VERSION : 0.1
// Master sequencing for automatic operation
   VAR_INPUT
      RST : Bool;   // Sequence reset
   END_VAR
   VAR_OUTPUT
      RNG : Bool;   // Sequence running
   END_VAR
   VAR
      CRNT_STEP : Int;
      STEP_001 : "500_SEQ_STEP";
      STEP_005 : "500_SEQ_STEP";
      STEP_010 : "500_SEQ_STEP";
      STEP_020 : "500_SEQ_STEP";
      STEP_030 : "500_SEQ_STEP";
      STEP_040 : "500_SEQ_STEP";
      STEP_050 : "500_SEQ_STEP";
      STEP_060 : "500_SEQ_STEP";
      STEP_070 : "500_SEQ_STEP";
      STEP_080 : "500_SEQ_STEP";
      STEP_090 : "500_SEQ_STEP";
      STEP_095 : "500_SEQ_STEP";
      STEP_100 : "500_SEQ_STEP";
      STEP_110 : "500_SEQ_STEP";
      STEP_120 : "500_SEQ_STEP";
      STEP_130 : "500_SEQ_STEP";
      STEP_140 : "500_SEQ_STEP";
      STEP_150 : "500_SEQ_STEP";
      STEP_160 : "500_SEQ_STEP";
      STEP_170 : "500_SEQ_STEP";
      STEP_180 : "500_SEQ_STEP";
      STEP_190 : "500_SEQ_STEP";
      STEP_200 : "500_SEQ_STEP";
      STEP_210 : "500_SEQ_STEP";
      STEP_220 : "500_SEQ_STEP";
      STEP_230 : "500_SEQ_STEP";
      STEP_240 : "500_SEQ_STEP";
      STEP_250 : "500_SEQ_STEP";
      STEP_260 : "500_SEQ_STEP";
      STEP_270 : "500_SEQ_STEP";
      STEP_300 : "500_SEQ_STEP";
      STEP_310 : "500_SEQ_STEP";
      STEP_320 : "500_SEQ_STEP";
      STEP_330 : "500_SEQ_STEP";
      STEP_340 : "500_SEQ_STEP";
      STEP_350 : "500_SEQ_STEP";
      STEP_360 : "500_SEQ_STEP";
      STEP_370 : "500_SEQ_STEP";
      STEP_380 : "500_SEQ_STEP";
      STEP_390 : "500_SEQ_STEP";
      STEP_400 : "500_SEQ_STEP";
      STEP_410 : "500_SEQ_STEP";
      STEP_420 : "500_SEQ_STEP";
      STEP_430 : "500_SEQ_STEP";
      STEP_440 : "500_SEQ_STEP";
      STEP_450 : "500_SEQ_STEP";
      STEP_460 : "500_SEQ_STEP";
      STEP_470 : "500_SEQ_STEP";
      STEP_480 : "500_SEQ_STEP";
      STEP_490 : "500_SEQ_STEP";
      STEP_500 : "500_SEQ_STEP";
      STEP_510 : "500_SEQ_STEP";
      STEP_520 : "500_SEQ_STEP";
      STEP_525 : "500_SEQ_STEP";
      STEP_530 : "500_SEQ_STEP";
      STEP_540 : "500_SEQ_STEP";
      STEP_550 : "500_SEQ_STEP";
      STEP_560 : "500_SEQ_STEP";
      STEP_570 : "500_SEQ_STEP";
   END_VAR
   VAR_TEMP   // added for the SCL form of the ladder/FBD networks
      _w1 : Bool;
   END_VAR
BEGIN

REGION Network 1: Auto Initiated or Reset = Set Step to 0
   // Going into automatic or sequence reset resets the sequence
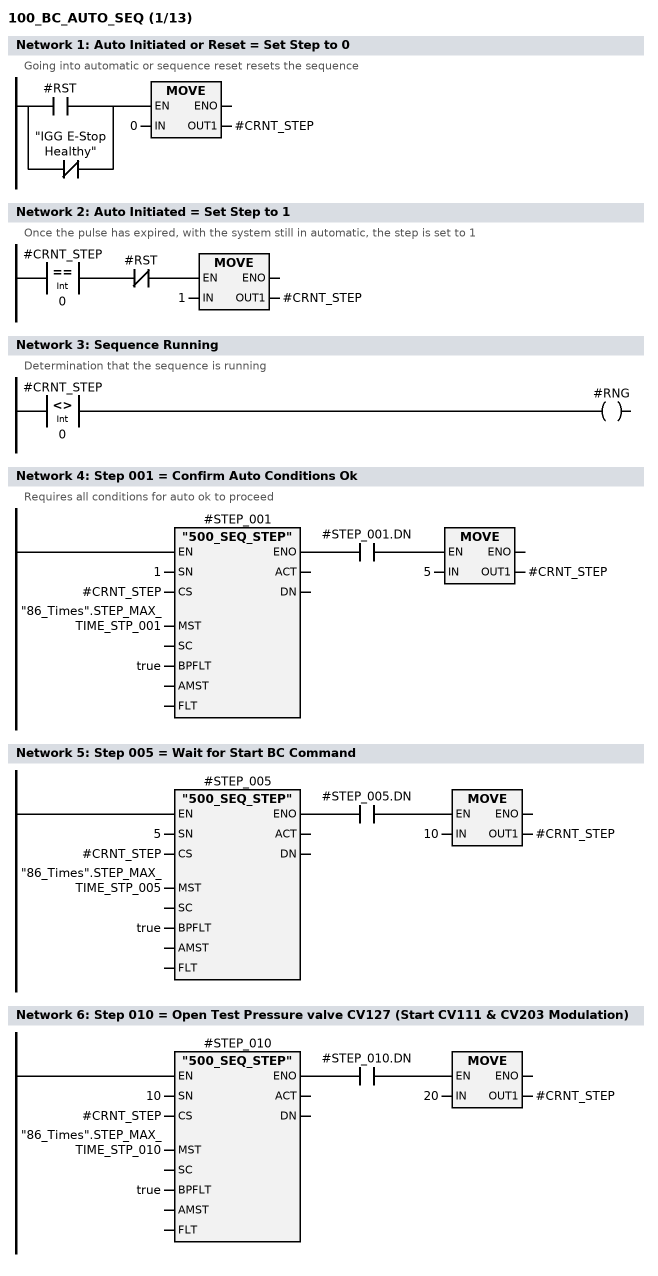
   RUNG wire#powerrail
      Contact( #RST )
      wire#w1
      Move(in := 0, out1 => #CRNT_STEP)
   END_RUNG
   RUNG wire#powerrail
      I_Contact( "IGG E-Stop Healthy" )
   END_RUNG wire#w1
   // the same network as SCL:
   IF #RST OR NOT "IGG E-Stop Healthy" THEN #CRNT_STEP := 0; END_IF;
END_REGION

REGION Network 2: Auto Initiated = Set Step to 1
   // Once the pulse has expired, with the system still in automatic, the step is set to 1
   RUNG wire#powerrail
      { S7_Templates := "SrcType := Int" } EQ_Contact(in1 := #CRNT_STEP, in2 := 0)
      I_Contact( #RST )
      Move(in := 1, out1 => #CRNT_STEP)
   END_RUNG
   // the same network as SCL:
   IF (#CRNT_STEP = 0) AND NOT #RST THEN #CRNT_STEP := 1; END_IF;
END_REGION

REGION Network 3: Sequence Running
   // Determination that the sequence is running
   RUNG wire#powerrail
      { S7_Templates := "SrcType := Int" } NE_Contact(in1 := #CRNT_STEP, in2 := 0)
      Coil( #RNG )
   END_RUNG
   // the same network as SCL:
   #RNG := #CRNT_STEP <> 0;
END_REGION

REGION Network 4: Step 001 = Confirm Auto Conditions Ok
   // Requires all conditions for auto ok to proceed
   RUNG wire#powerrail
      #STEP_001(SN := 1, CS := #CRNT_STEP, MST := "86_Times".STEP_MAX_TIME_STP_001, SC :=, BPFLT := true, AMST :=, FLT :=, ACT =>, DN =>)
      Contact( #STEP_001.DN )
      Move(in := 5, out1 => #CRNT_STEP)
   END_RUNG
   // the same network as SCL:
   #STEP_001(SN := 1, CS := #CRNT_STEP, MST := "86_Times".STEP_MAX_TIME_STP_001, BPFLT := true, ENO => #_w1);   // "500_SEQ_STEP"
   IF #_w1 AND #STEP_001.DN THEN #CRNT_STEP := 5; END_IF;
END_REGION

REGION Network 5: Step 005 = Wait for Start BC Command
   RUNG wire#powerrail
      #STEP_005(SN := 5, CS := #CRNT_STEP, MST := "86_Times".STEP_MAX_TIME_STP_005, SC :=, BPFLT := true, AMST :=, FLT :=, ACT =>, DN =>)
      Contact( #STEP_005.DN )
      Move(in := 10, out1 => #CRNT_STEP)
   END_RUNG
   // the same network as SCL:
   #STEP_005(SN := 5, CS := #CRNT_STEP, MST := "86_Times".STEP_MAX_TIME_STP_005, BPFLT := true, ENO => #_w1);   // "500_SEQ_STEP"
   IF #_w1 AND #STEP_005.DN THEN #CRNT_STEP := 10; END_IF;
END_REGION

REGION Network 6: Step 010 = Open Test Pressure valve CV127 (Start CV111 & CV203 Modulation)
   RUNG wire#powerrail
      #STEP_010(SN := 10, CS := #CRNT_STEP, MST := "86_Times".STEP_MAX_TIME_STP_010, SC :=, BPFLT := true, AMST :=, FLT :=, ACT =>, DN =>)
      Contact( #STEP_010.DN )
      Move(in := 20, out1 => #CRNT_STEP)
   END_RUNG
   // the same network as SCL:
   #STEP_010(SN := 10, CS := #CRNT_STEP, MST := "86_Times".STEP_MAX_TIME_STP_010, BPFLT := true, ENO => #_w1);   // "500_SEQ_STEP"
   IF #_w1 AND #STEP_010.DN THEN #CRNT_STEP := 20; END_IF;
END_REGION

REGION Network 7: Step 020 = Check Pressure PS101
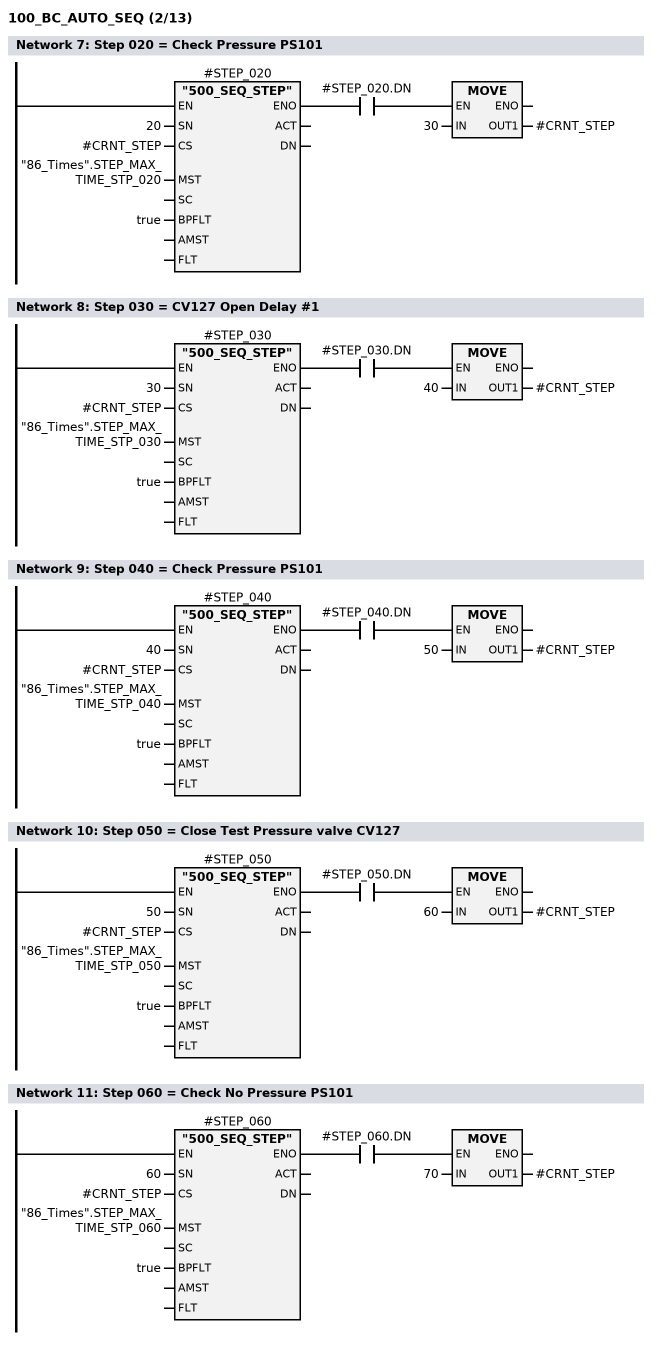
   RUNG wire#powerrail
      #STEP_020(SN := 20, CS := #CRNT_STEP, MST := "86_Times".STEP_MAX_TIME_STP_020, SC :=, BPFLT := true, AMST :=, FLT :=, ACT =>, DN =>)
      Contact( #STEP_020.DN )
      Move(in := 30, out1 => #CRNT_STEP)
   END_RUNG
   // the same network as SCL:
   #STEP_020(SN := 20, CS := #CRNT_STEP, MST := "86_Times".STEP_MAX_TIME_STP_020, BPFLT := true, ENO => #_w1);   // "500_SEQ_STEP"
   IF #_w1 AND #STEP_020.DN THEN #CRNT_STEP := 30; END_IF;
END_REGION

REGION Network 8: Step 030 = CV127 Open Delay #1
   RUNG wire#powerrail
      #STEP_030(SN := 30, CS := #CRNT_STEP, MST := "86_Times".STEP_MAX_TIME_STP_030, SC :=, BPFLT := true, AMST :=, FLT :=, ACT =>, DN =>)
      Contact( #STEP_030.DN )
      Move(in := 40, out1 => #CRNT_STEP)
   END_RUNG
   // the same network as SCL:
   #STEP_030(SN := 30, CS := #CRNT_STEP, MST := "86_Times".STEP_MAX_TIME_STP_030, BPFLT := true, ENO => #_w1);   // "500_SEQ_STEP"
   IF #_w1 AND #STEP_030.DN THEN #CRNT_STEP := 40; END_IF;
END_REGION

REGION Network 9: Step 040 = Check Pressure PS101
   RUNG wire#powerrail
      #STEP_040(SN := 40, CS := #CRNT_STEP, MST := "86_Times".STEP_MAX_TIME_STP_040, SC :=, BPFLT := true, AMST :=, FLT :=, ACT =>, DN =>)
      Contact( #STEP_040.DN )
      Move(in := 50, out1 => #CRNT_STEP)
   END_RUNG
   // the same network as SCL:
   #STEP_040(SN := 40, CS := #CRNT_STEP, MST := "86_Times".STEP_MAX_TIME_STP_040, BPFLT := true, ENO => #_w1);   // "500_SEQ_STEP"
   IF #_w1 AND #STEP_040.DN THEN #CRNT_STEP := 50; END_IF;
END_REGION

REGION Network 10: Step 050 = Close Test Pressure valve CV127
   RUNG wire#powerrail
      #STEP_050(SN := 50, CS := #CRNT_STEP, MST := "86_Times".STEP_MAX_TIME_STP_050, SC :=, BPFLT := true, AMST :=, FLT :=, ACT =>, DN =>)
      Contact( #STEP_050.DN )
      Move(in := 60, out1 => #CRNT_STEP)
   END_RUNG
   // the same network as SCL:
   #STEP_050(SN := 50, CS := #CRNT_STEP, MST := "86_Times".STEP_MAX_TIME_STP_050, BPFLT := true, ENO => #_w1);   // "500_SEQ_STEP"
   IF #_w1 AND #STEP_050.DN THEN #CRNT_STEP := 60; END_IF;
END_REGION

REGION Network 11: Step 060 = Check No Pressure PS101
   RUNG wire#powerrail
      #STEP_060(SN := 60, CS := #CRNT_STEP, MST := "86_Times".STEP_MAX_TIME_STP_060, SC :=, BPFLT := true, AMST :=, FLT :=, ACT =>, DN =>)
      Contact( #STEP_060.DN )
      Move(in := 70, out1 => #CRNT_STEP)
   END_RUNG
   // the same network as SCL:
   #STEP_060(SN := 60, CS := #CRNT_STEP, MST := "86_Times".STEP_MAX_TIME_STP_060, BPFLT := true, ENO => #_w1);   // "500_SEQ_STEP"
   IF #_w1 AND #STEP_060.DN THEN #CRNT_STEP := 70; END_IF;
END_REGION

REGION Network 12: Step 070 = CV127 Closed Delay
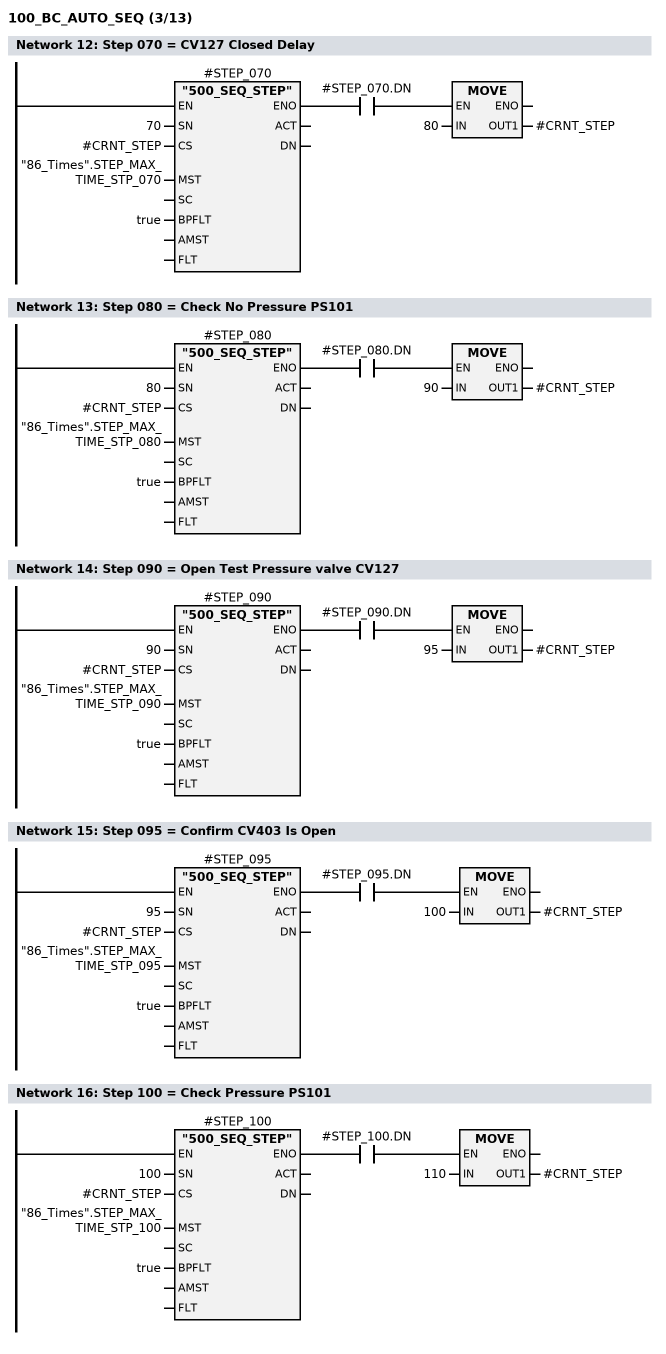
   RUNG wire#powerrail
      #STEP_070(SN := 70, CS := #CRNT_STEP, MST := "86_Times".STEP_MAX_TIME_STP_070, SC :=, BPFLT := true, AMST :=, FLT :=, ACT =>, DN =>)
      Contact( #STEP_070.DN )
      Move(in := 80, out1 => #CRNT_STEP)
   END_RUNG
   // the same network as SCL:
   #STEP_070(SN := 70, CS := #CRNT_STEP, MST := "86_Times".STEP_MAX_TIME_STP_070, BPFLT := true, ENO => #_w1);   // "500_SEQ_STEP"
   IF #_w1 AND #STEP_070.DN THEN #CRNT_STEP := 80; END_IF;
END_REGION

REGION Network 13: Step 080 = Check No Pressure PS101
   RUNG wire#powerrail
      #STEP_080(SN := 80, CS := #CRNT_STEP, MST := "86_Times".STEP_MAX_TIME_STP_080, SC :=, BPFLT := true, AMST :=, FLT :=, ACT =>, DN =>)
      Contact( #STEP_080.DN )
      Move(in := 90, out1 => #CRNT_STEP)
   END_RUNG
   // the same network as SCL:
   #STEP_080(SN := 80, CS := #CRNT_STEP, MST := "86_Times".STEP_MAX_TIME_STP_080, BPFLT := true, ENO => #_w1);   // "500_SEQ_STEP"
   IF #_w1 AND #STEP_080.DN THEN #CRNT_STEP := 90; END_IF;
END_REGION

REGION Network 14: Step 090 = Open Test Pressure valve CV127
   RUNG wire#powerrail
      #STEP_090(SN := 90, CS := #CRNT_STEP, MST := "86_Times".STEP_MAX_TIME_STP_090, SC :=, BPFLT := true, AMST :=, FLT :=, ACT =>, DN =>)
      Contact( #STEP_090.DN )
      Move(in := 95, out1 => #CRNT_STEP)
   END_RUNG
   // the same network as SCL:
   #STEP_090(SN := 90, CS := #CRNT_STEP, MST := "86_Times".STEP_MAX_TIME_STP_090, BPFLT := true, ENO => #_w1);   // "500_SEQ_STEP"
   IF #_w1 AND #STEP_090.DN THEN #CRNT_STEP := 95; END_IF;
END_REGION

REGION Network 15: Step 095 = Confirm CV403 Is Open
   RUNG wire#powerrail
      #STEP_095(SN := 95, CS := #CRNT_STEP, MST := "86_Times".STEP_MAX_TIME_STP_095, SC :=, BPFLT := true, AMST :=, FLT :=, ACT =>, DN =>)
      Contact( #STEP_095.DN )
      Move(in := 100, out1 => #CRNT_STEP)
   END_RUNG
   // the same network as SCL:
   #STEP_095(SN := 95, CS := #CRNT_STEP, MST := "86_Times".STEP_MAX_TIME_STP_095, BPFLT := true, ENO => #_w1);   // "500_SEQ_STEP"
   IF #_w1 AND #STEP_095.DN THEN #CRNT_STEP := 100; END_IF;
END_REGION

REGION Network 16: Step 100 = Check Pressure PS101
   RUNG wire#powerrail
      #STEP_100(SN := 100, CS := #CRNT_STEP, MST := "86_Times".STEP_MAX_TIME_STP_100, SC :=, BPFLT := true, AMST :=, FLT :=, ACT =>, DN =>)
      Contact( #STEP_100.DN )
      Move(in := 110, out1 => #CRNT_STEP)
   END_RUNG
   // the same network as SCL:
   #STEP_100(SN := 100, CS := #CRNT_STEP, MST := "86_Times".STEP_MAX_TIME_STP_100, BPFLT := true, ENO => #_w1);   // "500_SEQ_STEP"
   IF #_w1 AND #STEP_100.DN THEN #CRNT_STEP := 110; END_IF;
END_REGION

REGION Network 17: Step110 = CV127 Open Delay #2
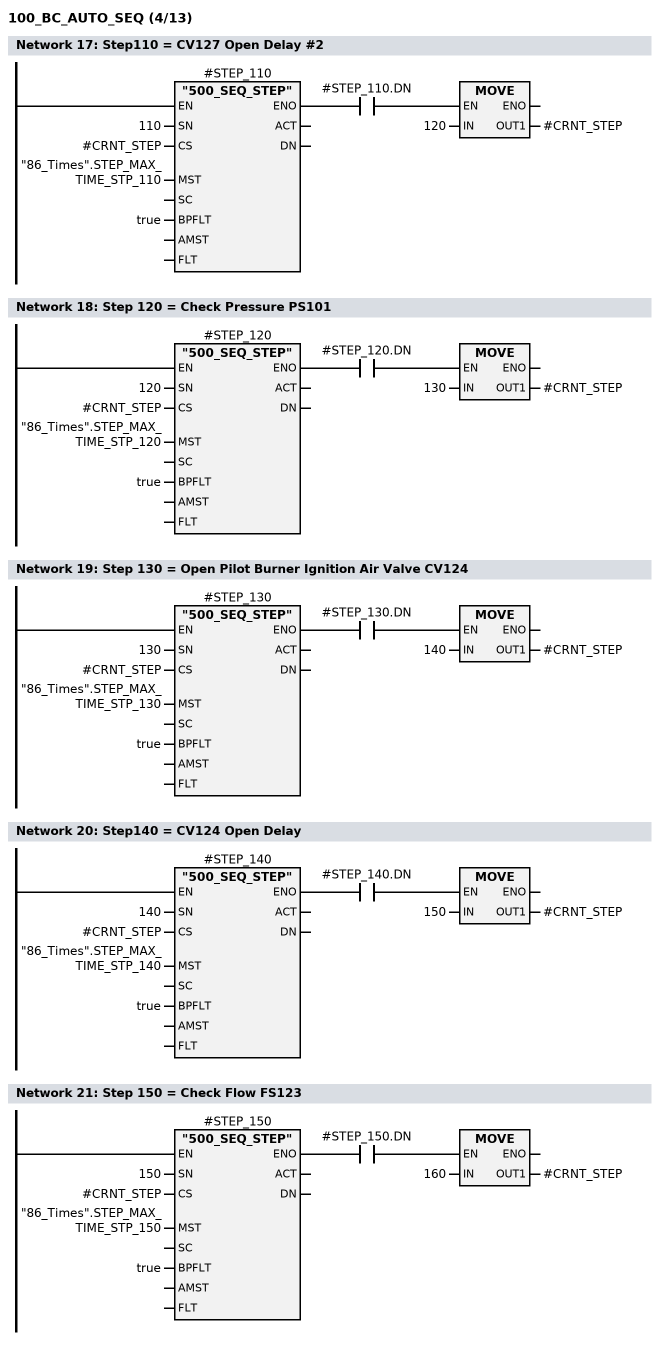
   RUNG wire#powerrail
      #STEP_110(SN := 110, CS := #CRNT_STEP, MST := "86_Times".STEP_MAX_TIME_STP_110, SC :=, BPFLT := true, AMST :=, FLT :=, ACT =>, DN =>)
      Contact( #STEP_110.DN )
      Move(in := 120, out1 => #CRNT_STEP)
   END_RUNG
   // the same network as SCL:
   #STEP_110(SN := 110, CS := #CRNT_STEP, MST := "86_Times".STEP_MAX_TIME_STP_110, BPFLT := true, ENO => #_w1);   // "500_SEQ_STEP"
   IF #_w1 AND #STEP_110.DN THEN #CRNT_STEP := 120; END_IF;
END_REGION

REGION Network 18: Step 120 = Check Pressure PS101
   RUNG wire#powerrail
      #STEP_120(SN := 120, CS := #CRNT_STEP, MST := "86_Times".STEP_MAX_TIME_STP_120, SC :=, BPFLT := true, AMST :=, FLT :=, ACT =>, DN =>)
      Contact( #STEP_120.DN )
      Move(in := 130, out1 => #CRNT_STEP)
   END_RUNG
   // the same network as SCL:
   #STEP_120(SN := 120, CS := #CRNT_STEP, MST := "86_Times".STEP_MAX_TIME_STP_120, BPFLT := true, ENO => #_w1);   // "500_SEQ_STEP"
   IF #_w1 AND #STEP_120.DN THEN #CRNT_STEP := 130; END_IF;
END_REGION

REGION Network 19: Step 130 = Open Pilot Burner Ignition Air Valve CV124
   RUNG wire#powerrail
      #STEP_130(SN := 130, CS := #CRNT_STEP, MST := "86_Times".STEP_MAX_TIME_STP_130, SC :=, BPFLT := true, AMST :=, FLT :=, ACT =>, DN =>)
      Contact( #STEP_130.DN )
      Move(in := 140, out1 => #CRNT_STEP)
   END_RUNG
   // the same network as SCL:
   #STEP_130(SN := 130, CS := #CRNT_STEP, MST := "86_Times".STEP_MAX_TIME_STP_130, BPFLT := true, ENO => #_w1);   // "500_SEQ_STEP"
   IF #_w1 AND #STEP_130.DN THEN #CRNT_STEP := 140; END_IF;
END_REGION

REGION Network 20: Step140 = CV124 Open Delay
   RUNG wire#powerrail
      #STEP_140(SN := 140, CS := #CRNT_STEP, MST := "86_Times".STEP_MAX_TIME_STP_140, SC :=, BPFLT := true, AMST :=, FLT :=, ACT =>, DN =>)
      Contact( #STEP_140.DN )
      Move(in := 150, out1 => #CRNT_STEP)
   END_RUNG
   // the same network as SCL:
   #STEP_140(SN := 140, CS := #CRNT_STEP, MST := "86_Times".STEP_MAX_TIME_STP_140, BPFLT := true, ENO => #_w1);   // "500_SEQ_STEP"
   IF #_w1 AND #STEP_140.DN THEN #CRNT_STEP := 150; END_IF;
END_REGION

REGION Network 21: Step 150 = Check Flow FS123
   RUNG wire#powerrail
      #STEP_150(SN := 150, CS := #CRNT_STEP, MST := "86_Times".STEP_MAX_TIME_STP_150, SC :=, BPFLT := true, AMST :=, FLT :=, ACT =>, DN =>)
      Contact( #STEP_150.DN )
      Move(in := 160, out1 => #CRNT_STEP)
   END_RUNG
   // the same network as SCL:
   #STEP_150(SN := 150, CS := #CRNT_STEP, MST := "86_Times".STEP_MAX_TIME_STP_150, BPFLT := true, ENO => #_w1);   // "500_SEQ_STEP"
   IF #_w1 AND #STEP_150.DN THEN #CRNT_STEP := 160; END_IF;
END_REGION

REGION Network 22: Step 160 = Pilot Flame Ignition Sequence
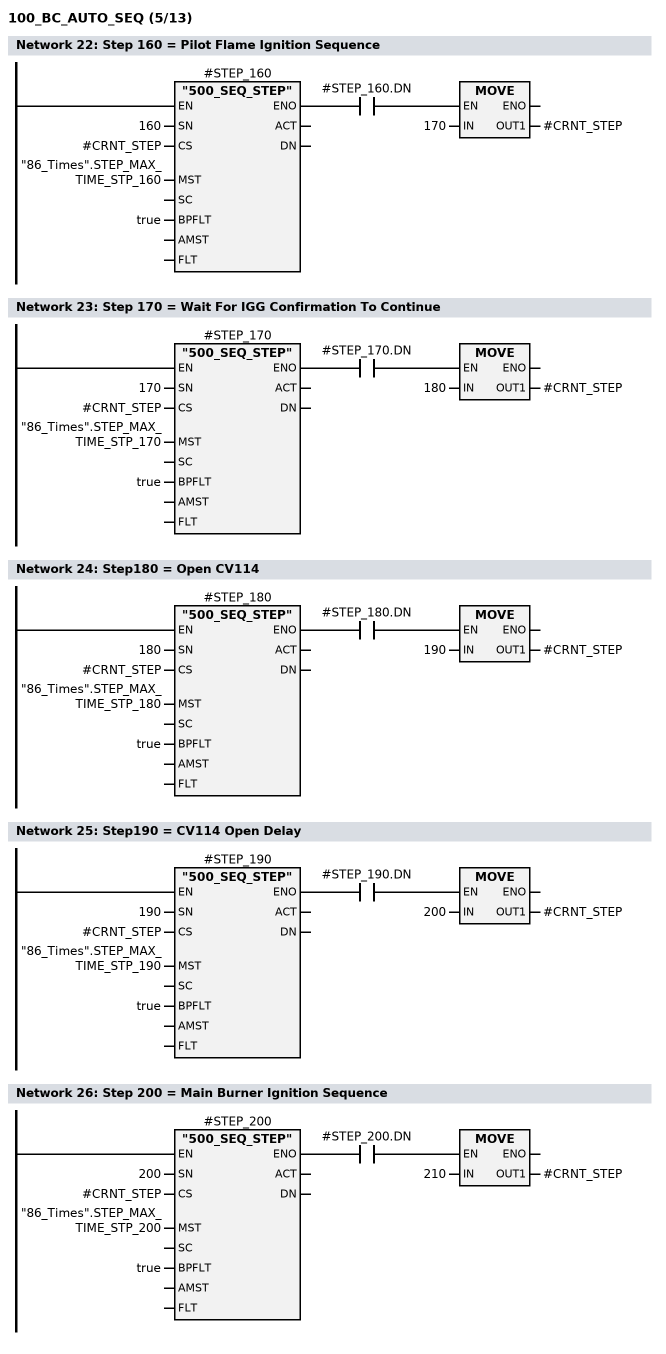
   RUNG wire#powerrail
      #STEP_160(SN := 160, CS := #CRNT_STEP, MST := "86_Times".STEP_MAX_TIME_STP_160, SC :=, BPFLT := true, AMST :=, FLT :=, ACT =>, DN =>)
      Contact( #STEP_160.DN )
      Move(in := 170, out1 => #CRNT_STEP)
   END_RUNG
   // the same network as SCL:
   #STEP_160(SN := 160, CS := #CRNT_STEP, MST := "86_Times".STEP_MAX_TIME_STP_160, BPFLT := true, ENO => #_w1);   // "500_SEQ_STEP"
   IF #_w1 AND #STEP_160.DN THEN #CRNT_STEP := 170; END_IF;
END_REGION

REGION Network 23: Step 170 = Wait For IGG Confirmation To Continue
   RUNG wire#powerrail
      #STEP_170(SN := 170, CS := #CRNT_STEP, MST := "86_Times".STEP_MAX_TIME_STP_170, SC :=, BPFLT := true, AMST :=, FLT :=, ACT =>, DN =>)
      Contact( #STEP_170.DN )
      Move(in := 180, out1 => #CRNT_STEP)
   END_RUNG
   // the same network as SCL:
   #STEP_170(SN := 170, CS := #CRNT_STEP, MST := "86_Times".STEP_MAX_TIME_STP_170, BPFLT := true, ENO => #_w1);   // "500_SEQ_STEP"
   IF #_w1 AND #STEP_170.DN THEN #CRNT_STEP := 180; END_IF;
END_REGION

REGION Network 24: Step180 = Open CV114
   RUNG wire#powerrail
      #STEP_180(SN := 180, CS := #CRNT_STEP, MST := "86_Times".STEP_MAX_TIME_STP_180, SC :=, BPFLT := true, AMST :=, FLT :=, ACT =>, DN =>)
      Contact( #STEP_180.DN )
      Move(in := 190, out1 => #CRNT_STEP)
   END_RUNG
   // the same network as SCL:
   #STEP_180(SN := 180, CS := #CRNT_STEP, MST := "86_Times".STEP_MAX_TIME_STP_180, BPFLT := true, ENO => #_w1);   // "500_SEQ_STEP"
   IF #_w1 AND #STEP_180.DN THEN #CRNT_STEP := 190; END_IF;
END_REGION

REGION Network 25: Step190 = CV114 Open Delay
   RUNG wire#powerrail
      #STEP_190(SN := 190, CS := #CRNT_STEP, MST := "86_Times".STEP_MAX_TIME_STP_190, SC :=, BPFLT := true, AMST :=, FLT :=, ACT =>, DN =>)
      Contact( #STEP_190.DN )
      Move(in := 200, out1 => #CRNT_STEP)
   END_RUNG
   // the same network as SCL:
   #STEP_190(SN := 190, CS := #CRNT_STEP, MST := "86_Times".STEP_MAX_TIME_STP_190, BPFLT := true, ENO => #_w1);   // "500_SEQ_STEP"
   IF #_w1 AND #STEP_190.DN THEN #CRNT_STEP := 200; END_IF;
END_REGION

REGION Network 26: Step 200 = Main Burner Ignition Sequence
   RUNG wire#powerrail
      #STEP_200(SN := 200, CS := #CRNT_STEP, MST := "86_Times".STEP_MAX_TIME_STP_200, SC :=, BPFLT := true, AMST :=, FLT :=, ACT =>, DN =>)
      Contact( #STEP_200.DN )
      Move(in := 210, out1 => #CRNT_STEP)
   END_RUNG
   // the same network as SCL:
   #STEP_200(SN := 200, CS := #CRNT_STEP, MST := "86_Times".STEP_MAX_TIME_STP_200, BPFLT := true, ENO => #_w1);   // "500_SEQ_STEP"
   IF #_w1 AND #STEP_200.DN THEN #CRNT_STEP := 210; END_IF;
END_REGION

REGION Network 27: Step 210 = Check Pressure PIT113
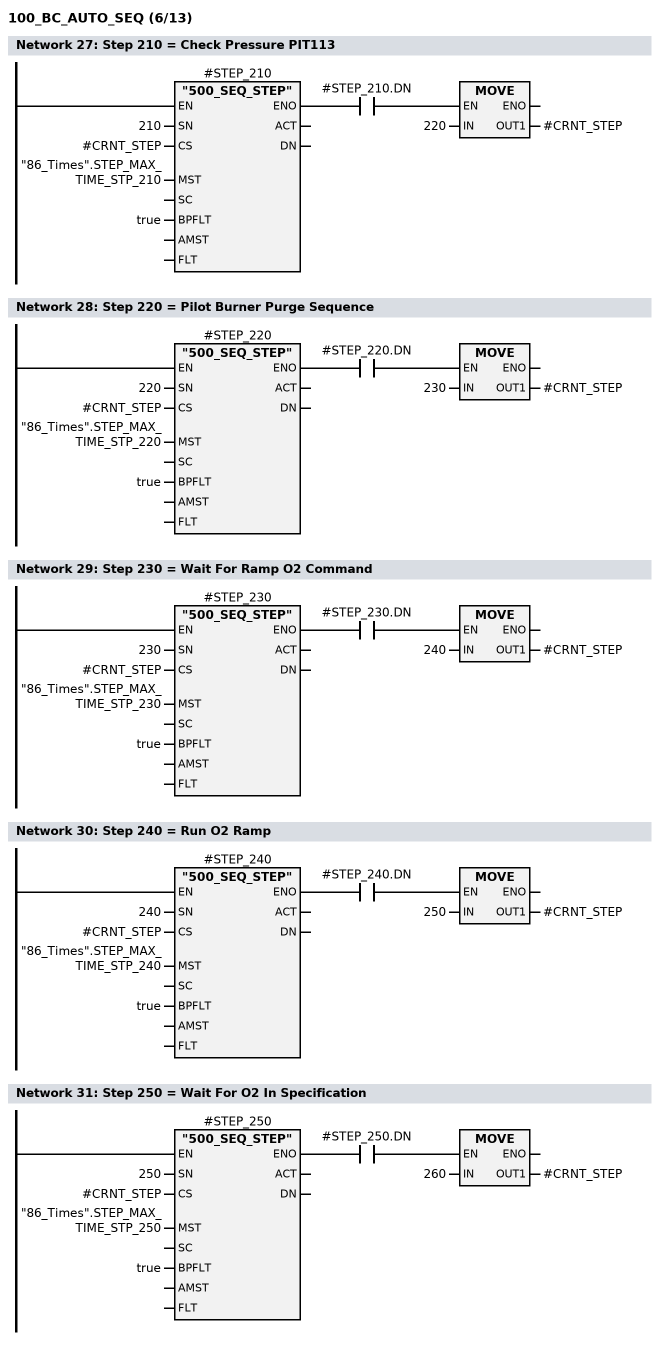
   RUNG wire#powerrail
      #STEP_210(SN := 210, CS := #CRNT_STEP, MST := "86_Times".STEP_MAX_TIME_STP_210, SC :=, BPFLT := true, AMST :=, FLT :=, ACT =>, DN =>)
      Contact( #STEP_210.DN )
      Move(in := 220, out1 => #CRNT_STEP)
   END_RUNG
   // the same network as SCL:
   #STEP_210(SN := 210, CS := #CRNT_STEP, MST := "86_Times".STEP_MAX_TIME_STP_210, BPFLT := true, ENO => #_w1);   // "500_SEQ_STEP"
   IF #_w1 AND #STEP_210.DN THEN #CRNT_STEP := 220; END_IF;
END_REGION

REGION Network 28: Step 220 = Pilot Burner Purge Sequence
   RUNG wire#powerrail
      #STEP_220(SN := 220, CS := #CRNT_STEP, MST := "86_Times".STEP_MAX_TIME_STP_220, SC :=, BPFLT := true, AMST :=, FLT :=, ACT =>, DN =>)
      Contact( #STEP_220.DN )
      Move(in := 230, out1 => #CRNT_STEP)
   END_RUNG
   // the same network as SCL:
   #STEP_220(SN := 220, CS := #CRNT_STEP, MST := "86_Times".STEP_MAX_TIME_STP_220, BPFLT := true, ENO => #_w1);   // "500_SEQ_STEP"
   IF #_w1 AND #STEP_220.DN THEN #CRNT_STEP := 230; END_IF;
END_REGION

REGION Network 29: Step 230 = Wait For Ramp O2 Command
   RUNG wire#powerrail
      #STEP_230(SN := 230, CS := #CRNT_STEP, MST := "86_Times".STEP_MAX_TIME_STP_230, SC :=, BPFLT := true, AMST :=, FLT :=, ACT =>, DN =>)
      Contact( #STEP_230.DN )
      Move(in := 240, out1 => #CRNT_STEP)
   END_RUNG
   // the same network as SCL:
   #STEP_230(SN := 230, CS := #CRNT_STEP, MST := "86_Times".STEP_MAX_TIME_STP_230, BPFLT := true, ENO => #_w1);   // "500_SEQ_STEP"
   IF #_w1 AND #STEP_230.DN THEN #CRNT_STEP := 240; END_IF;
END_REGION

REGION Network 30: Step 240 = Run O2 Ramp
   RUNG wire#powerrail
      #STEP_240(SN := 240, CS := #CRNT_STEP, MST := "86_Times".STEP_MAX_TIME_STP_240, SC :=, BPFLT := true, AMST :=, FLT :=, ACT =>, DN =>)
      Contact( #STEP_240.DN )
      Move(in := 250, out1 => #CRNT_STEP)
   END_RUNG
   // the same network as SCL:
   #STEP_240(SN := 240, CS := #CRNT_STEP, MST := "86_Times".STEP_MAX_TIME_STP_240, BPFLT := true, ENO => #_w1);   // "500_SEQ_STEP"
   IF #_w1 AND #STEP_240.DN THEN #CRNT_STEP := 250; END_IF;
END_REGION

REGION Network 31: Step 250 = Wait For O2 In Specification
   RUNG wire#powerrail
      #STEP_250(SN := 250, CS := #CRNT_STEP, MST := "86_Times".STEP_MAX_TIME_STP_250, SC :=, BPFLT := true, AMST :=, FLT :=, ACT =>, DN =>)
      Contact( #STEP_250.DN )
      Move(in := 260, out1 => #CRNT_STEP)
   END_RUNG
   // the same network as SCL:
   #STEP_250(SN := 250, CS := #CRNT_STEP, MST := "86_Times".STEP_MAX_TIME_STP_250, BPFLT := true, ENO => #_w1);   // "500_SEQ_STEP"
   IF #_w1 AND #STEP_250.DN THEN #CRNT_STEP := 260; END_IF;
END_REGION

REGION Network 32: Step 260 = Write O2 Within Specification Status To IGG
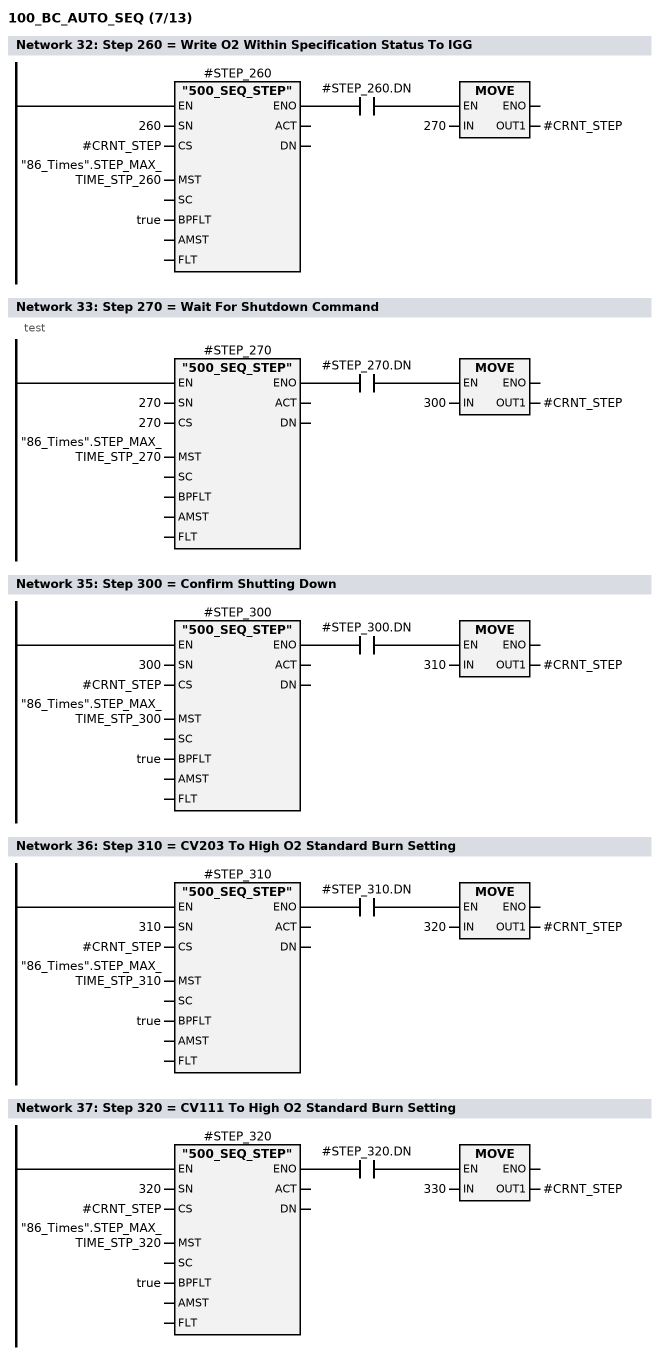
   RUNG wire#powerrail
      #STEP_260(SN := 260, CS := #CRNT_STEP, MST := "86_Times".STEP_MAX_TIME_STP_260, SC :=, BPFLT := true, AMST :=, FLT :=, ACT =>, DN =>)
      Contact( #STEP_260.DN )
      Move(in := 270, out1 => #CRNT_STEP)
   END_RUNG
   // the same network as SCL:
   #STEP_260(SN := 260, CS := #CRNT_STEP, MST := "86_Times".STEP_MAX_TIME_STP_260, BPFLT := true, ENO => #_w1);   // "500_SEQ_STEP"
   IF #_w1 AND #STEP_260.DN THEN #CRNT_STEP := 270; END_IF;
END_REGION

REGION Network 33: Step 270 = Wait For Shutdown Command
   // test
   RUNG wire#powerrail
      #STEP_270(SN := 270, CS := 270, MST := "86_Times".STEP_MAX_TIME_STP_270, SC :=, BPFLT :=, AMST :=, FLT :=, ACT =>, DN =>)
      Contact( #STEP_270.DN )
      Move(in := 300, out1 => #CRNT_STEP)
   END_RUNG
   // the same network as SCL:
   #STEP_270(SN := 270, CS := 270, MST := "86_Times".STEP_MAX_TIME_STP_270, ENO => #_w1);   // "500_SEQ_STEP"
   IF #_w1 AND #STEP_270.DN THEN #CRNT_STEP := 300; END_IF;
END_REGION

REGION Network 35: Step 300 = Confirm Shutting Down
   RUNG wire#powerrail
      #STEP_300(SN := 300, CS := #CRNT_STEP, MST := "86_Times".STEP_MAX_TIME_STP_300, SC :=, BPFLT := true, AMST :=, FLT :=, ACT =>, DN =>)
      Contact( #STEP_300.DN )
      Move(in := 310, out1 => #CRNT_STEP)
   END_RUNG
   // the same network as SCL:
   #STEP_300(SN := 300, CS := #CRNT_STEP, MST := "86_Times".STEP_MAX_TIME_STP_300, BPFLT := true, ENO => #_w1);   // "500_SEQ_STEP"
   IF #_w1 AND #STEP_300.DN THEN #CRNT_STEP := 310; END_IF;
END_REGION

REGION Network 36: Step 310 = CV203 To High O2 Standard Burn Setting
   RUNG wire#powerrail
      #STEP_310(SN := 310, CS := #CRNT_STEP, MST := "86_Times".STEP_MAX_TIME_STP_310, SC :=, BPFLT := true, AMST :=, FLT :=, ACT =>, DN =>)
      Contact( #STEP_310.DN )
      Move(in := 320, out1 => #CRNT_STEP)
   END_RUNG
   // the same network as SCL:
   #STEP_310(SN := 310, CS := #CRNT_STEP, MST := "86_Times".STEP_MAX_TIME_STP_310, BPFLT := true, ENO => #_w1);   // "500_SEQ_STEP"
   IF #_w1 AND #STEP_310.DN THEN #CRNT_STEP := 320; END_IF;
END_REGION

REGION Network 37: Step 320 = CV111 To High O2 Standard Burn Setting
   RUNG wire#powerrail
      #STEP_320(SN := 320, CS := #CRNT_STEP, MST := "86_Times".STEP_MAX_TIME_STP_320, SC :=, BPFLT := true, AMST :=, FLT :=, ACT =>, DN =>)
      Contact( #STEP_320.DN )
      Move(in := 330, out1 => #CRNT_STEP)
   END_RUNG
   // the same network as SCL:
   #STEP_320(SN := 320, CS := #CRNT_STEP, MST := "86_Times".STEP_MAX_TIME_STP_320, BPFLT := true, ENO => #_w1);   // "500_SEQ_STEP"
   IF #_w1 AND #STEP_320.DN THEN #CRNT_STEP := 330; END_IF;
END_REGION

REGION Network 38: Step 330 = Modulation Stopped Confirmation To IGG
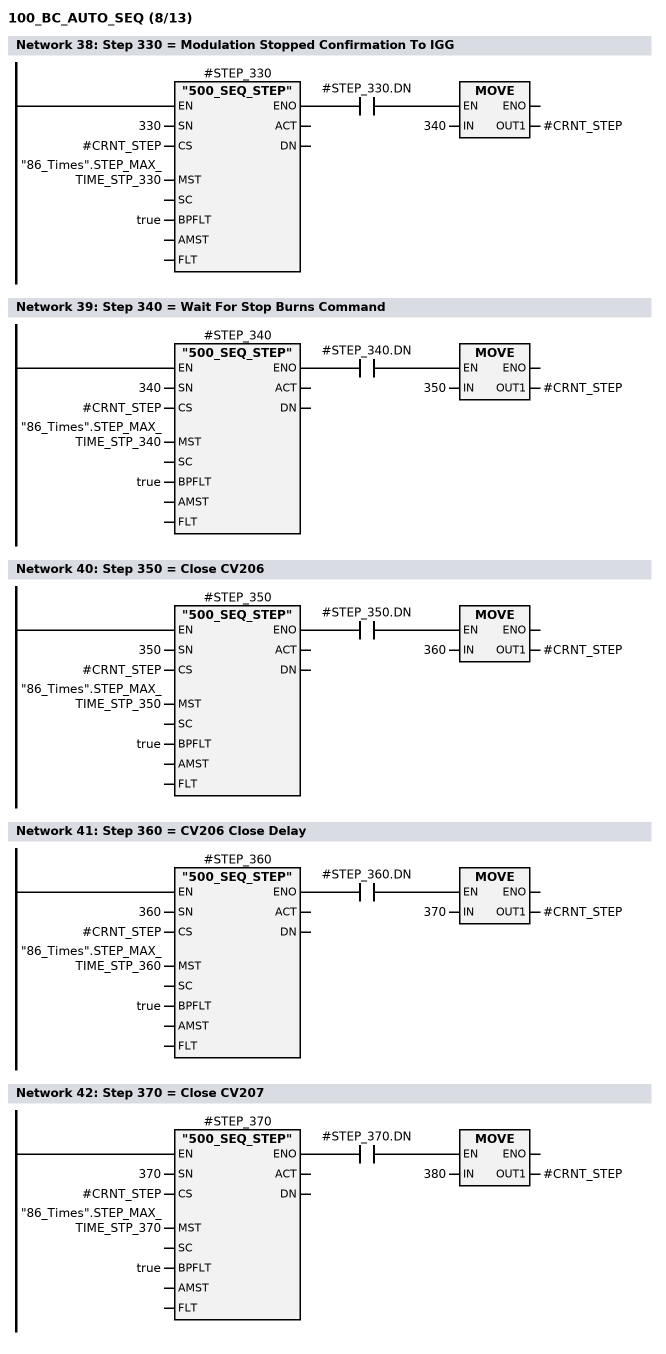
   RUNG wire#powerrail
      #STEP_330(SN := 330, CS := #CRNT_STEP, MST := "86_Times".STEP_MAX_TIME_STP_330, SC :=, BPFLT := true, AMST :=, FLT :=, ACT =>, DN =>)
      Contact( #STEP_330.DN )
      Move(in := 340, out1 => #CRNT_STEP)
   END_RUNG
   // the same network as SCL:
   #STEP_330(SN := 330, CS := #CRNT_STEP, MST := "86_Times".STEP_MAX_TIME_STP_330, BPFLT := true, ENO => #_w1);   // "500_SEQ_STEP"
   IF #_w1 AND #STEP_330.DN THEN #CRNT_STEP := 340; END_IF;
END_REGION

REGION Network 39: Step 340 = Wait For Stop Burns Command
   RUNG wire#powerrail
      #STEP_340(SN := 340, CS := #CRNT_STEP, MST := "86_Times".STEP_MAX_TIME_STP_340, SC :=, BPFLT := true, AMST :=, FLT :=, ACT =>, DN =>)
      Contact( #STEP_340.DN )
      Move(in := 350, out1 => #CRNT_STEP)
   END_RUNG
   // the same network as SCL:
   #STEP_340(SN := 340, CS := #CRNT_STEP, MST := "86_Times".STEP_MAX_TIME_STP_340, BPFLT := true, ENO => #_w1);   // "500_SEQ_STEP"
   IF #_w1 AND #STEP_340.DN THEN #CRNT_STEP := 350; END_IF;
END_REGION

REGION Network 40: Step 350 = Close CV206
   RUNG wire#powerrail
      #STEP_350(SN := 350, CS := #CRNT_STEP, MST := "86_Times".STEP_MAX_TIME_STP_350, SC :=, BPFLT := true, AMST :=, FLT :=, ACT =>, DN =>)
      Contact( #STEP_350.DN )
      Move(in := 360, out1 => #CRNT_STEP)
   END_RUNG
   // the same network as SCL:
   #STEP_350(SN := 350, CS := #CRNT_STEP, MST := "86_Times".STEP_MAX_TIME_STP_350, BPFLT := true, ENO => #_w1);   // "500_SEQ_STEP"
   IF #_w1 AND #STEP_350.DN THEN #CRNT_STEP := 360; END_IF;
END_REGION

REGION Network 41: Step 360 = CV206 Close Delay
   RUNG wire#powerrail
      #STEP_360(SN := 360, CS := #CRNT_STEP, MST := "86_Times".STEP_MAX_TIME_STP_360, SC :=, BPFLT := true, AMST :=, FLT :=, ACT =>, DN =>)
      Contact( #STEP_360.DN )
      Move(in := 370, out1 => #CRNT_STEP)
   END_RUNG
   // the same network as SCL:
   #STEP_360(SN := 360, CS := #CRNT_STEP, MST := "86_Times".STEP_MAX_TIME_STP_360, BPFLT := true, ENO => #_w1);   // "500_SEQ_STEP"
   IF #_w1 AND #STEP_360.DN THEN #CRNT_STEP := 370; END_IF;
END_REGION

REGION Network 42: Step 370 = Close CV207
   RUNG wire#powerrail
      #STEP_370(SN := 370, CS := #CRNT_STEP, MST := "86_Times".STEP_MAX_TIME_STP_370, SC :=, BPFLT := true, AMST :=, FLT :=, ACT =>, DN =>)
      Contact( #STEP_370.DN )
      Move(in := 380, out1 => #CRNT_STEP)
   END_RUNG
   // the same network as SCL:
   #STEP_370(SN := 370, CS := #CRNT_STEP, MST := "86_Times".STEP_MAX_TIME_STP_370, BPFLT := true, ENO => #_w1);   // "500_SEQ_STEP"
   IF #_w1 AND #STEP_370.DN THEN #CRNT_STEP := 380; END_IF;
END_REGION

REGION Network 43: Step 380 = CV207 Close Delay
